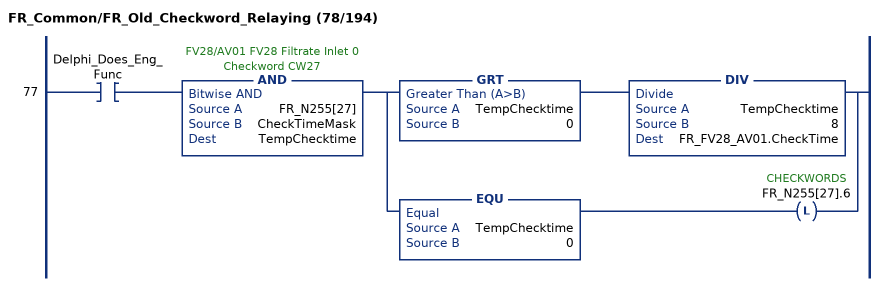
   77: XIC(Delphi_Does_Eng_Func)AND(FR_N255[27],CheckTimeMask,TempChecktime)[GRT(TempChecktime,0) DIV(TempChecktime,8,FR_FV28_AV01.CheckTime) ,EQU(TempChecktime,0) OTL(FR_N255[27].6) ];
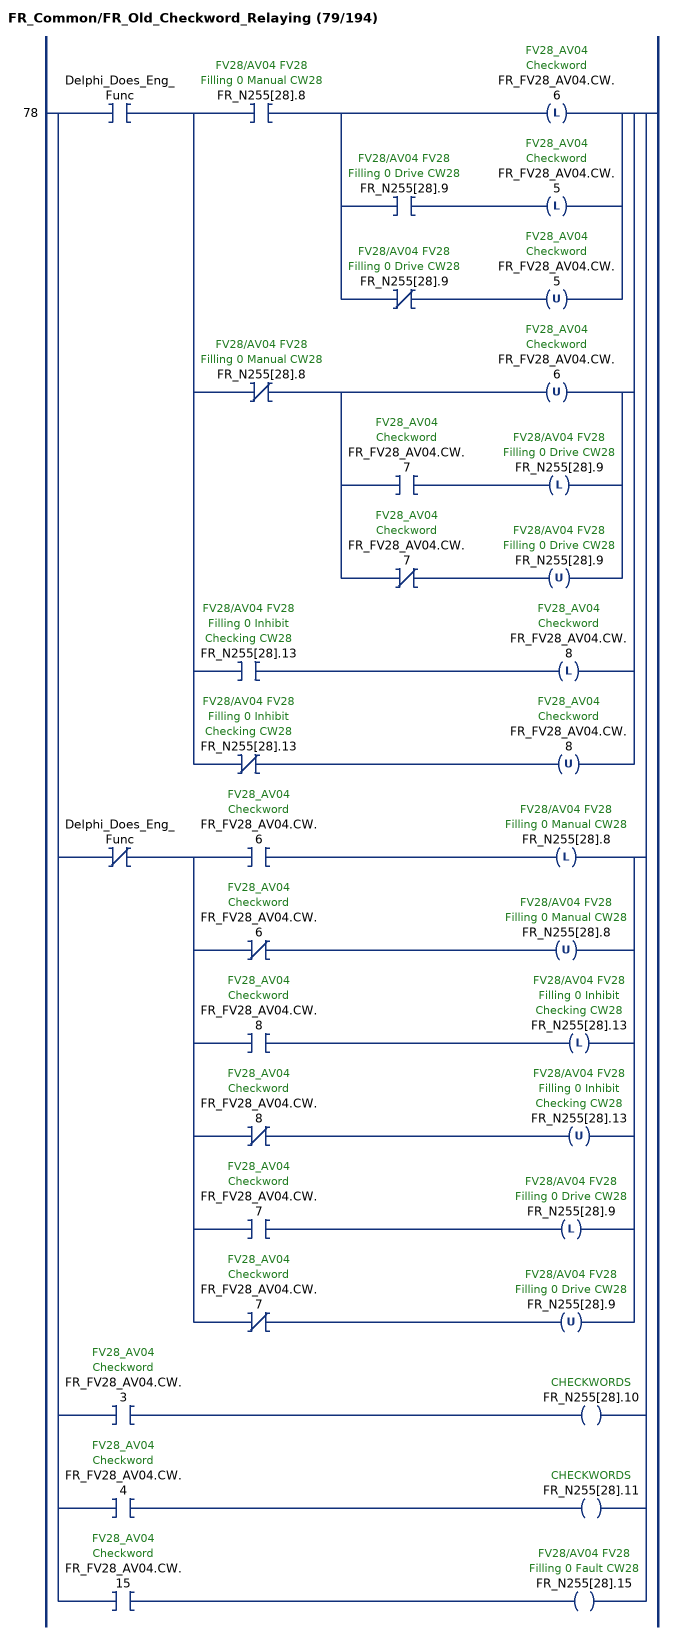
   78: [XIC(Delphi_Does_Eng_Func) [[XIC(FR_N255[28].8) [OTL(FR_FV28_AV04.CW.6) ,XIC(FR_N255[28].9) OTL(FR_FV28_AV04.CW.5) ,XIO(FR_N255[28].9) OTU(FR_FV28_AV04.CW.5) ] ,XIO(FR_N255[28].8) [OTU(FR_FV28_AV04.CW.6) ,[XIC(FR_FV28_AV04.CW.7) OTL(FR_N255[28].9) ,XIO(FR_FV28_AV04.CW.7) OTU(FR_N255[28].9) ] ] ] ,[XIC(FR_N255[28].13) OTL(FR_FV28_AV04.CW.8) ,XIO(FR_N255[28].13) OTU(FR_FV28_AV04.CW.8) ] ] ,XIO(Delphi_Does_Eng_Func) [[XIC(FR_FV28_AV04.CW.6) OTL(FR_N255[28].8) ,XIO(FR_FV28_AV04.CW.6) OTU(FR_N255[28].8) ] ,[XIC(FR_FV28_AV04.CW.8) OTL(FR_N255[28].13) ,XIO(FR_FV28_AV04.CW.8) OTU(FR_N255[28].13) ] ,[XIC(FR_FV28_AV04.CW.7) OTL(FR_N255[28].9) ,XIO(FR_FV28_AV04.CW.7) OTU(FR_N255[28].9) ] ] ,XIC(FR_FV28_AV04.CW.3) OTE(FR_N255[28].10) ,XIC(FR_FV28_AV04.CW.4) OTE(FR_N255[28].11) ,XIC(FR_FV28_AV04.CW.15) OTE(FR_N255[28].15) ];
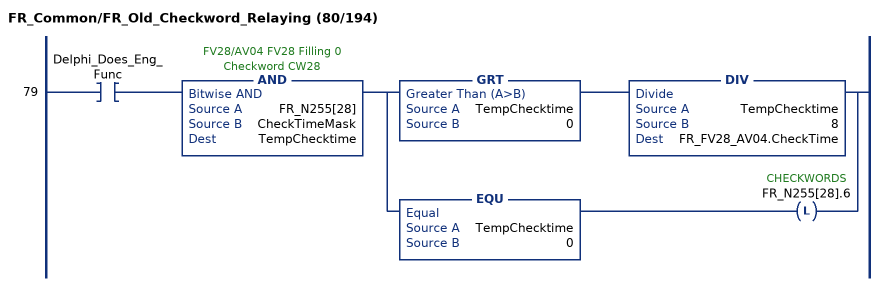
   79: XIC(Delphi_Does_Eng_Func)AND(FR_N255[28],CheckTimeMask,TempChecktime)[GRT(TempChecktime,0) DIV(TempChecktime,8,FR_FV28_AV04.CheckTime) ,EQU(TempChecktime,0) OTL(FR_N255[28].6) ];
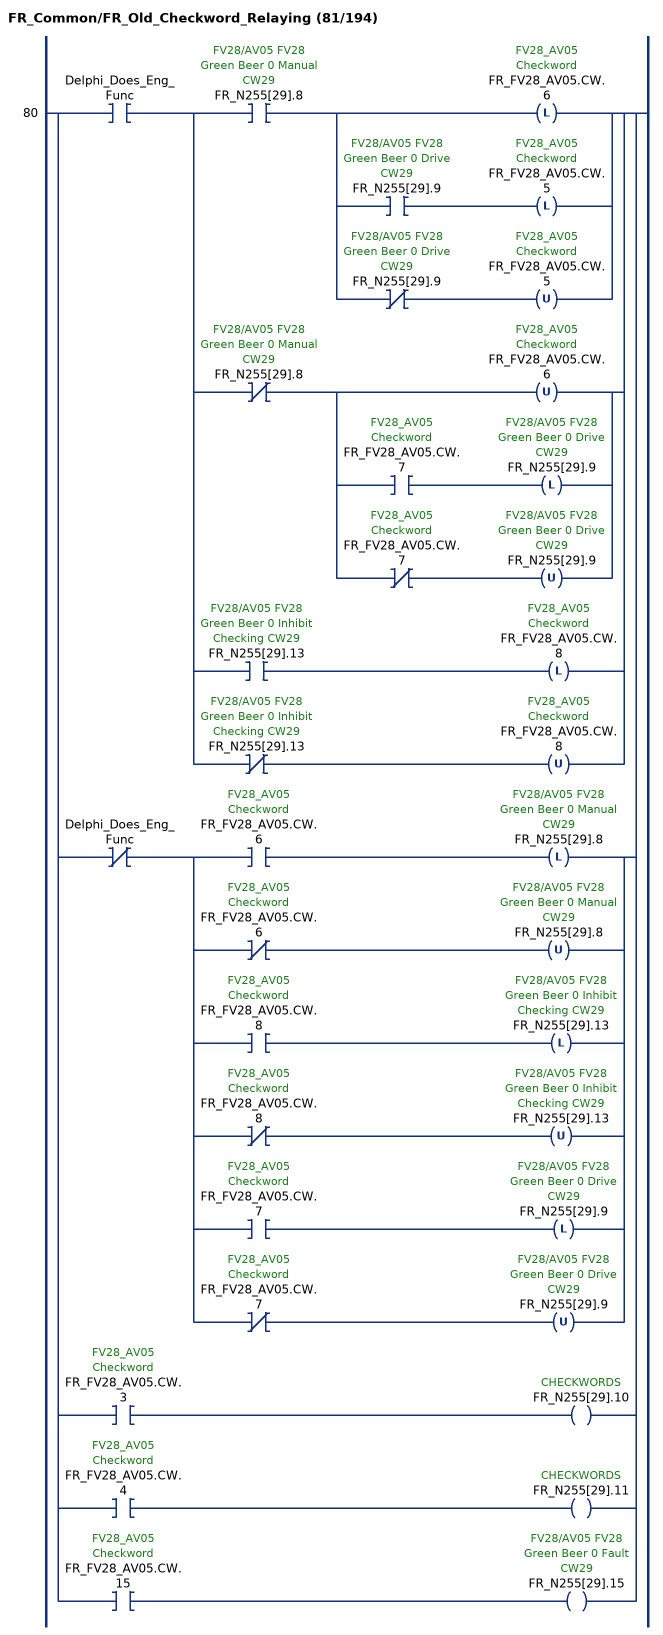
   80: [XIC(Delphi_Does_Eng_Func) [[XIC(FR_N255[29].8) [OTL(FR_FV28_AV05.CW.6) ,XIC(FR_N255[29].9) OTL(FR_FV28_AV05.CW.5) ,XIO(FR_N255[29].9) OTU(FR_FV28_AV05.CW.5) ] ,XIO(FR_N255[29].8) [OTU(FR_FV28_AV05.CW.6) ,[XIC(FR_FV28_AV05.CW.7) OTL(FR_N255[29].9) ,XIO(FR_FV28_AV05.CW.7) OTU(FR_N255[29].9) ] ] ] ,[XIC(FR_N255[29].13) OTL(FR_FV28_AV05.CW.8) ,XIO(FR_N255[29].13) OTU(FR_FV28_AV05.CW.8) ] ] ,XIO(Delphi_Does_Eng_Func) [[XIC(FR_FV28_AV05.CW.6) OTL(FR_N255[29].8) ,XIO(FR_FV28_AV05.CW.6) OTU(FR_N255[29].8) ] ,[XIC(FR_FV28_AV05.CW.8) OTL(FR_N255[29].13) ,XIO(FR_FV28_AV05.CW.8) OTU(FR_N255[29].13) ] ,[XIC(FR_FV28_AV05.CW.7) OTL(FR_N255[29].9) ,XIO(FR_FV28_AV05.CW.7) OTU(FR_N255[29].9) ] ] ,XIC(FR_FV28_AV05.CW.3) OTE(FR_N255[29].10) ,XIC(FR_FV28_AV05.CW.4) OTE(FR_N255[29].11) ,XIC(FR_FV28_AV05.CW.15) OTE(FR_N255[29].15) ];
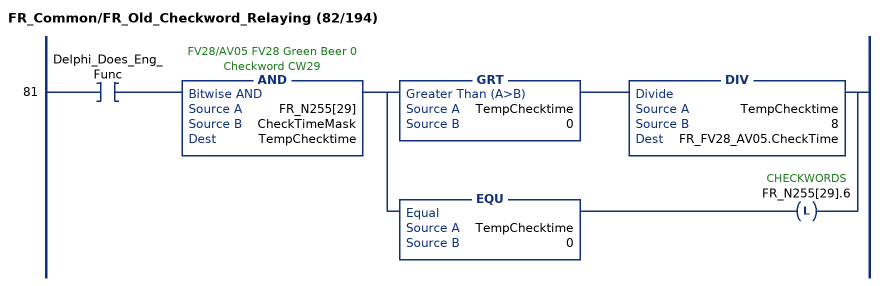
   81: XIC(Delphi_Does_Eng_Func)AND(FR_N255[29],CheckTimeMask,TempChecktime)[GRT(TempChecktime,0) DIV(TempChecktime,8,FR_FV28_AV05.CheckTime) ,EQU(TempChecktime,0) OTL(FR_N255[29].6) ];
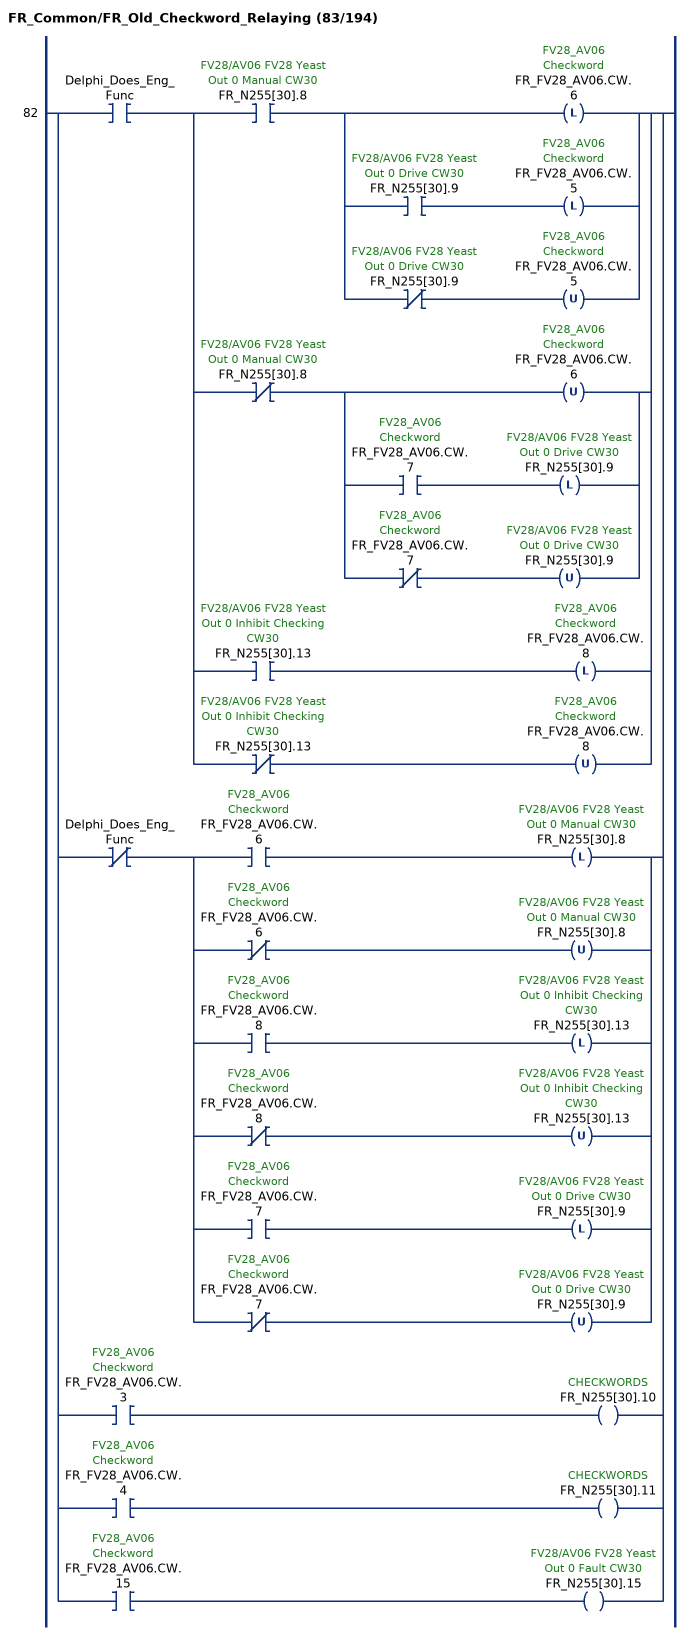
   82: [XIC(Delphi_Does_Eng_Func) [[XIC(FR_N255[30].8) [OTL(FR_FV28_AV06.CW.6) ,XIC(FR_N255[30].9) OTL(FR_FV28_AV06.CW.5) ,XIO(FR_N255[30].9) OTU(FR_FV28_AV06.CW.5) ] ,XIO(FR_N255[30].8) [OTU(FR_FV28_AV06.CW.6) ,[XIC(FR_FV28_AV06.CW.7) OTL(FR_N255[30].9) ,XIO(FR_FV28_AV06.CW.7) OTU(FR_N255[30].9) ] ] ] ,[XIC(FR_N255[30].13) OTL(FR_FV28_AV06.CW.8) ,XIO(FR_N255[30].13) OTU(FR_FV28_AV06.CW.8) ] ] ,XIO(Delphi_Does_Eng_Func) [[XIC(FR_FV28_AV06.CW.6) OTL(FR_N255[30].8) ,XIO(FR_FV28_AV06.CW.6) OTU(FR_N255[30].8) ] ,[XIC(FR_FV28_AV06.CW.8) OTL(FR_N255[30].13) ,XIO(FR_FV28_AV06.CW.8) OTU(FR_N255[30].13) ] ,[XIC(FR_FV28_AV06.CW.7) OTL(FR_N255[30].9) ,XIO(FR_FV28_AV06.CW.7) OTU(FR_N255[30].9) ] ] ,XIC(FR_FV28_AV06.CW.3) OTE(FR_N255[30].10) ,XIC(FR_FV28_AV06.CW.4) OTE(FR_N255[30].11) ,XIC(FR_FV28_AV06.CW.15) OTE(FR_N255[30].15) ];
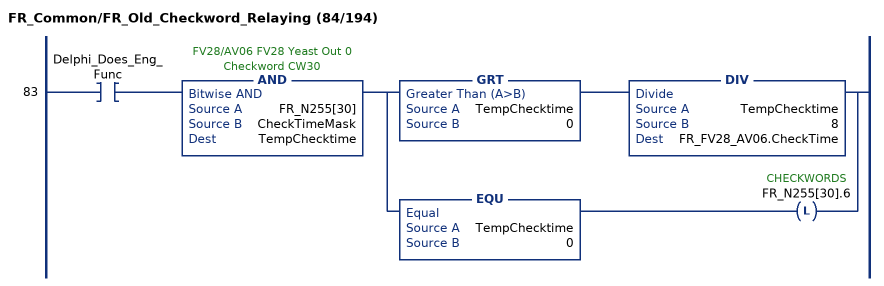
   83: XIC(Delphi_Does_Eng_Func)AND(FR_N255[30],CheckTimeMask,TempChecktime)[GRT(TempChecktime,0) DIV(TempChecktime,8,FR_FV28_AV06.CheckTime) ,EQU(TempChecktime,0) OTL(FR_N255[30].6) ];
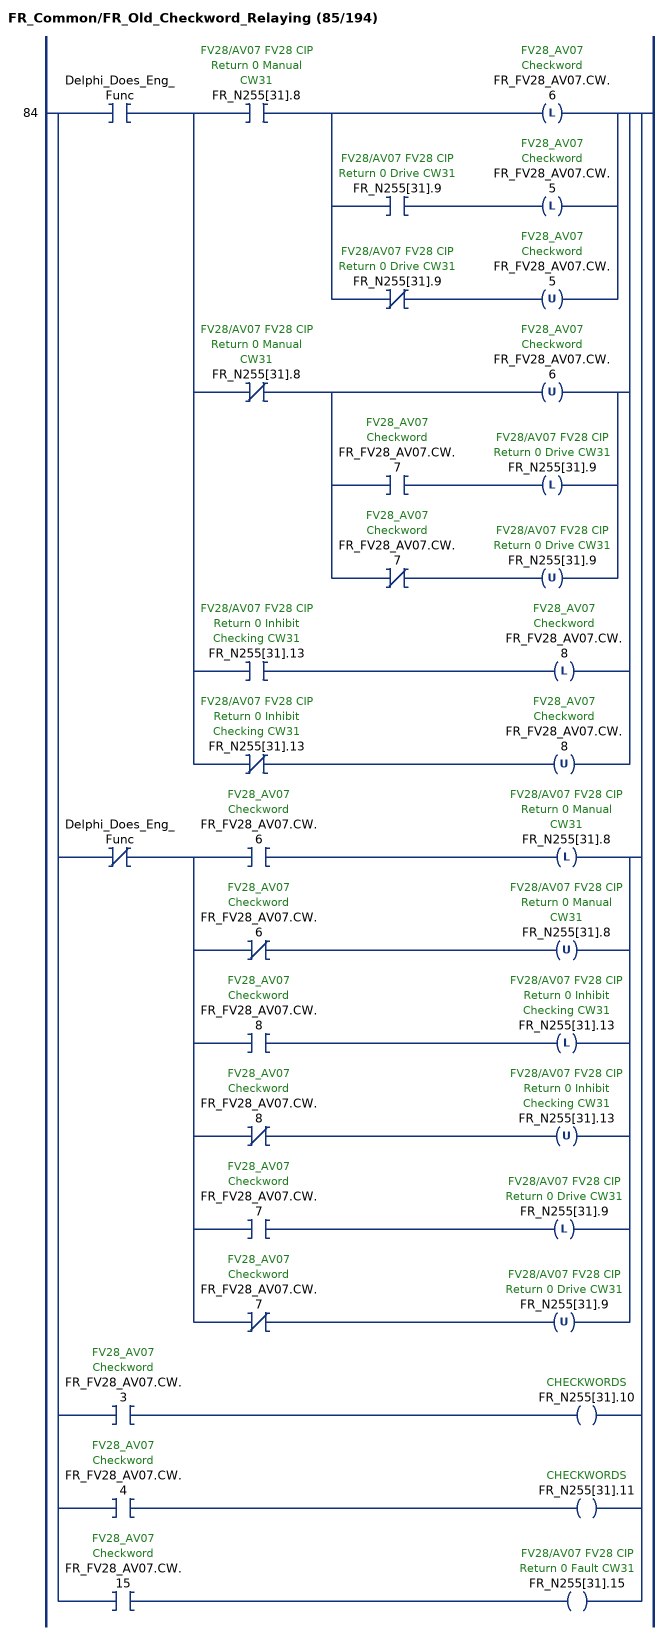
   84: [XIC(Delphi_Does_Eng_Func) [[XIC(FR_N255[31].8) [OTL(FR_FV28_AV07.CW.6) ,XIC(FR_N255[31].9) OTL(FR_FV28_AV07.CW.5) ,XIO(FR_N255[31].9) OTU(FR_FV28_AV07.CW.5) ] ,XIO(FR_N255[31].8) [OTU(FR_FV28_AV07.CW.6) ,[XIC(FR_FV28_AV07.CW.7) OTL(FR_N255[31].9) ,XIO(FR_FV28_AV07.CW.7) OTU(FR_N255[31].9) ] ] ] ,[XIC(FR_N255[31].13) OTL(FR_FV28_AV07.CW.8) ,XIO(FR_N255[31].13) OTU(FR_FV28_AV07.CW.8) ] ] ,XIO(Delphi_Does_Eng_Func) [[XIC(FR_FV28_AV07.CW.6) OTL(FR_N255[31].8) ,XIO(FR_FV28_AV07.CW.6) OTU(FR_N255[31].8) ] ,[XIC(FR_FV28_AV07.CW.8) OTL(FR_N255[31].13) ,XIO(FR_FV28_AV07.CW.8) OTU(FR_N255[31].13) ] ,[XIC(FR_FV28_AV07.CW.7) OTL(FR_N255[31].9) ,XIO(FR_FV28_AV07.CW.7) OTU(FR_N255[31].9) ] ] ,XIC(FR_FV28_AV07.CW.3) OTE(FR_N255[31].10) ,XIC(FR_FV28_AV07.CW.4) OTE(FR_N255[31].11) ,XIC(FR_FV28_AV07.CW.15) OTE(FR_N255[31].15) ];
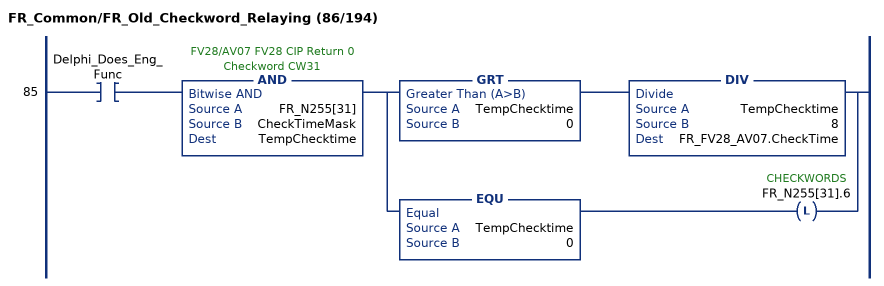
   85: XIC(Delphi_Does_Eng_Func)AND(FR_N255[31],CheckTimeMask,TempChecktime)[GRT(TempChecktime,0) DIV(TempChecktime,8,FR_FV28_AV07.CheckTime) ,EQU(TempChecktime,0) OTL(FR_N255[31].6) ];
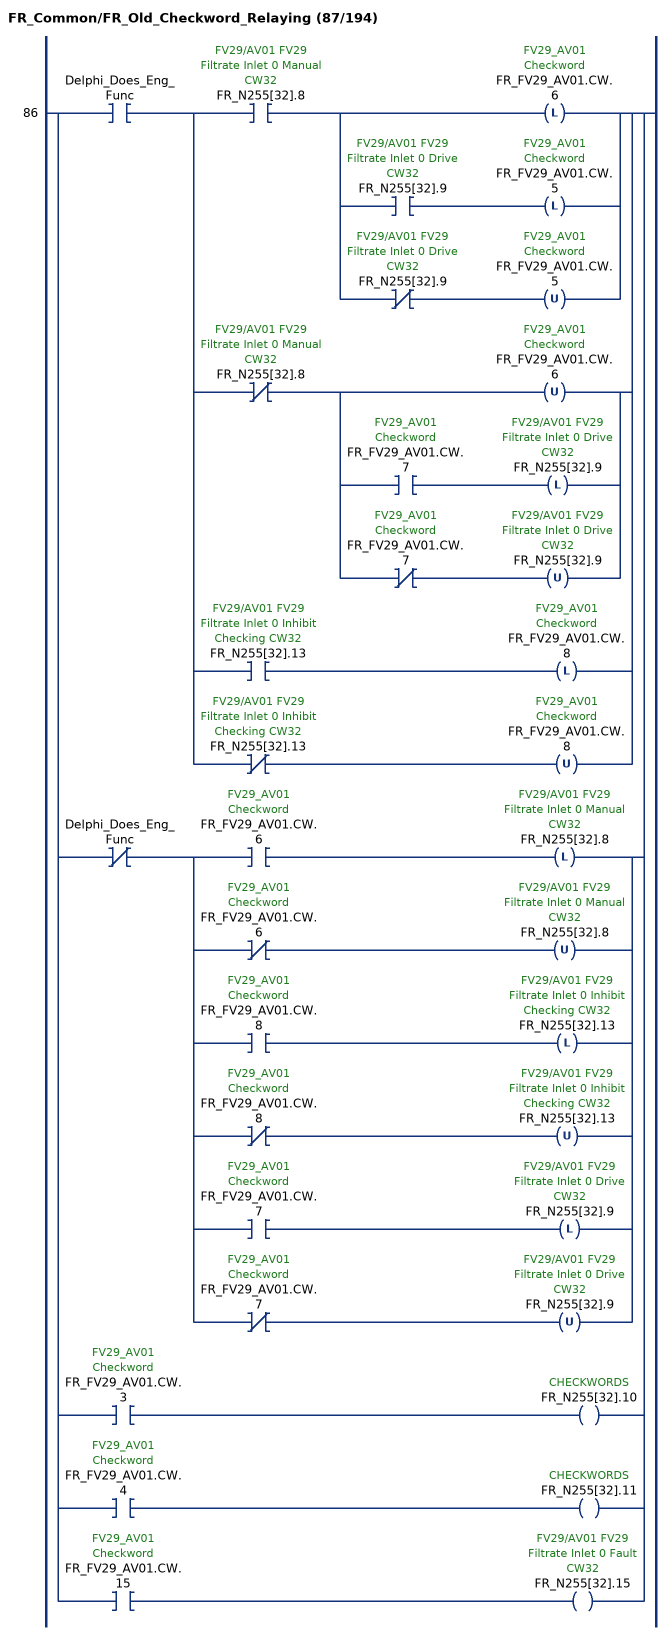
   86: [XIC(Delphi_Does_Eng_Func) [[XIC(FR_N255[32].8) [OTL(FR_FV29_AV01.CW.6) ,XIC(FR_N255[32].9) OTL(FR_FV29_AV01.CW.5) ,XIO(FR_N255[32].9) OTU(FR_FV29_AV01.CW.5) ] ,XIO(FR_N255[32].8) [OTU(FR_FV29_AV01.CW.6) ,[XIC(FR_FV29_AV01.CW.7) OTL(FR_N255[32].9) ,XIO(FR_FV29_AV01.CW.7) OTU(FR_N255[32].9) ] ] ] ,[XIC(FR_N255[32].13) OTL(FR_FV29_AV01.CW.8) ,XIO(FR_N255[32].13) OTU(FR_FV29_AV01.CW.8) ] ] ,XIO(Delphi_Does_Eng_Func) [[XIC(FR_FV29_AV01.CW.6) OTL(FR_N255[32].8) ,XIO(FR_FV29_AV01.CW.6) OTU(FR_N255[32].8) ] ,[XIC(FR_FV29_AV01.CW.8) OTL(FR_N255[32].13) ,XIO(FR_FV29_AV01.CW.8) OTU(FR_N255[32].13) ] ,[XIC(FR_FV29_AV01.CW.7) OTL(FR_N255[32].9) ,XIO(FR_FV29_AV01.CW.7) OTU(FR_N255[32].9) ] ] ,XIC(FR_FV29_AV01.CW.3) OTE(FR_N255[32].10) ,XIC(FR_FV29_AV01.CW.4) OTE(FR_N255[32].11) ,XIC(FR_FV29_AV01.CW.15) OTE(FR_N255[32].15) ];
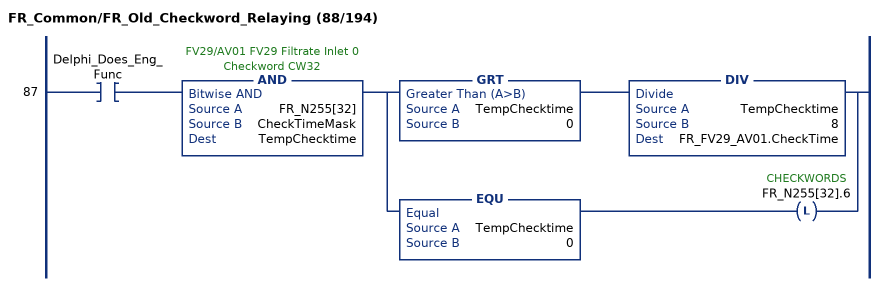
   87: XIC(Delphi_Does_Eng_Func)AND(FR_N255[32],CheckTimeMask,TempChecktime)[GRT(TempChecktime,0) DIV(TempChecktime,8,FR_FV29_AV01.CheckTime) ,EQU(TempChecktime,0) OTL(FR_N255[32].6) ];
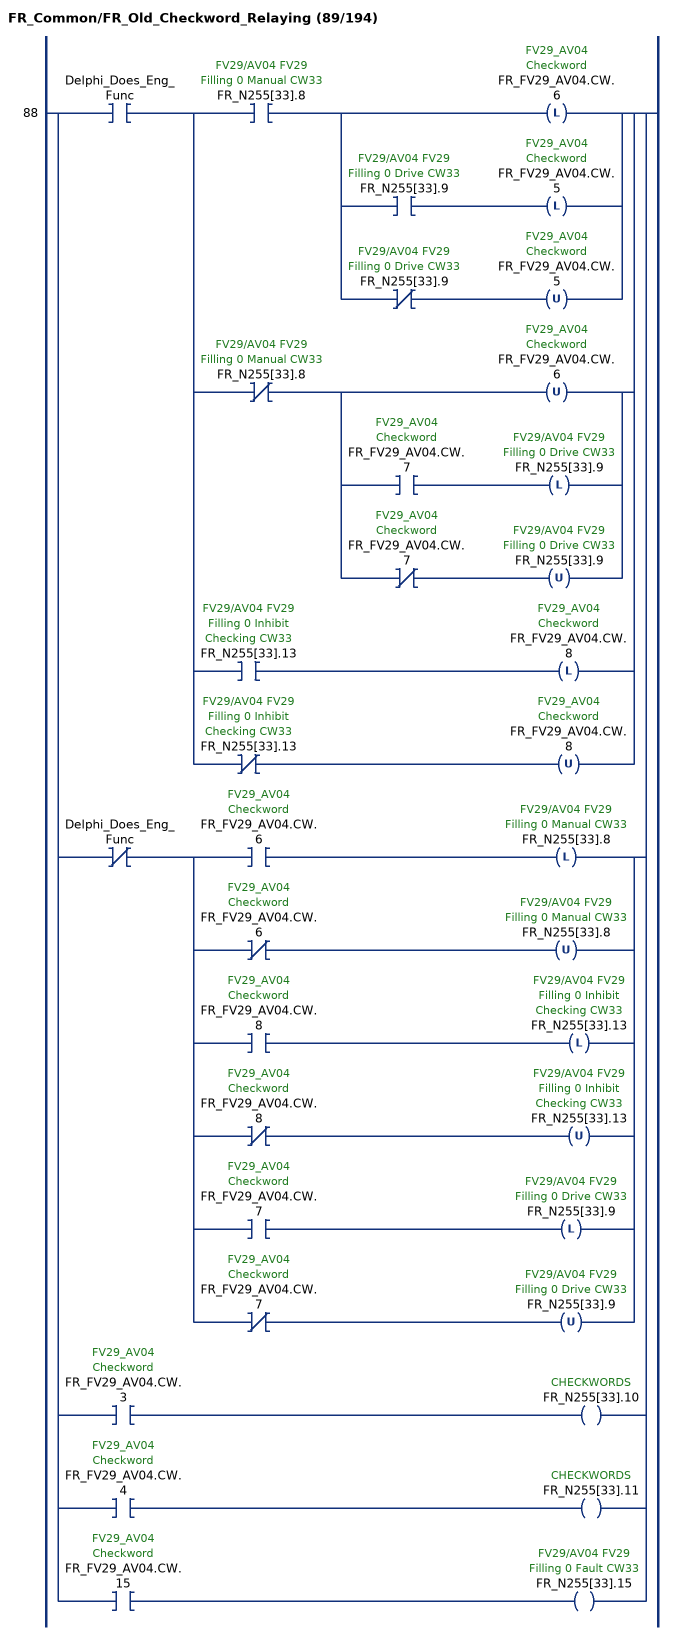
   88: [XIC(Delphi_Does_Eng_Func) [[XIC(FR_N255[33].8) [OTL(FR_FV29_AV04.CW.6) ,XIC(FR_N255[33].9) OTL(FR_FV29_AV04.CW.5) ,XIO(FR_N255[33].9) OTU(FR_FV29_AV04.CW.5) ] ,XIO(FR_N255[33].8) [OTU(FR_FV29_AV04.CW.6) ,[XIC(FR_FV29_AV04.CW.7) OTL(FR_N255[33].9) ,XIO(FR_FV29_AV04.CW.7) OTU(FR_N255[33].9) ] ] ] ,[XIC(FR_N255[33].13) OTL(FR_FV29_AV04.CW.8) ,XIO(FR_N255[33].13) OTU(FR_FV29_AV04.CW.8) ] ] ,XIO(Delphi_Does_Eng_Func) [[XIC(FR_FV29_AV04.CW.6) OTL(FR_N255[33].8) ,XIO(FR_FV29_AV04.CW.6) OTU(FR_N255[33].8) ] ,[XIC(FR_FV29_AV04.CW.8) OTL(FR_N255[33].13) ,XIO(FR_FV29_AV04.CW.8) OTU(FR_N255[33].13) ] ,[XIC(FR_FV29_AV04.CW.7) OTL(FR_N255[33].9) ,XIO(FR_FV29_AV04.CW.7) OTU(FR_N255[33].9) ] ] ,XIC(FR_FV29_AV04.CW.3) OTE(FR_N255[33].10) ,XIC(FR_FV29_AV04.CW.4) OTE(FR_N255[33].11) ,XIC(FR_FV29_AV04.CW.15) OTE(FR_N255[33].15) ];
